(* Logix 5000 project; controller _GigaDiscovery vendor 1 type 14 code 244 rev 35.11; software revision 35.03; part 11 of 23 *)
(* tags used below, declared in another part *)
   Emergencies_CL1 : DINT[14];
(* S_Alarms, continued *)

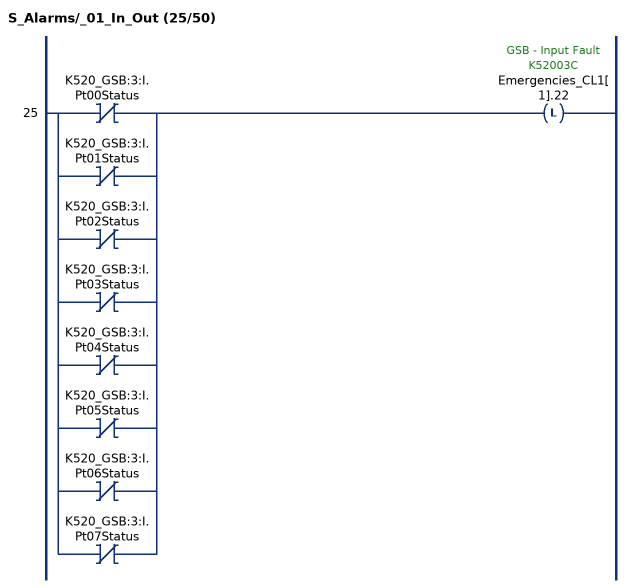
   [picture p185: S_Alarms/_01_In_Out rungs 25-25]
   25: [XIO(K520_GSB:3:I.Pt00Status) ,XIO(K520_GSB:3:I.Pt01Status) ,XIO(K520_GSB:3:I.Pt02Status) ,XIO(K520_GSB:3:I.Pt03Status) ,XIO(K520_GSB:3:I.Pt04Status) ,XIO(K520_GSB:3:I.Pt05Status) ,XIO(K520_GSB:3:I.Pt06Status) ,XIO(K520_GSB:3:I.Pt07Status) ]OTL(Emergencies_CL1[1].22);
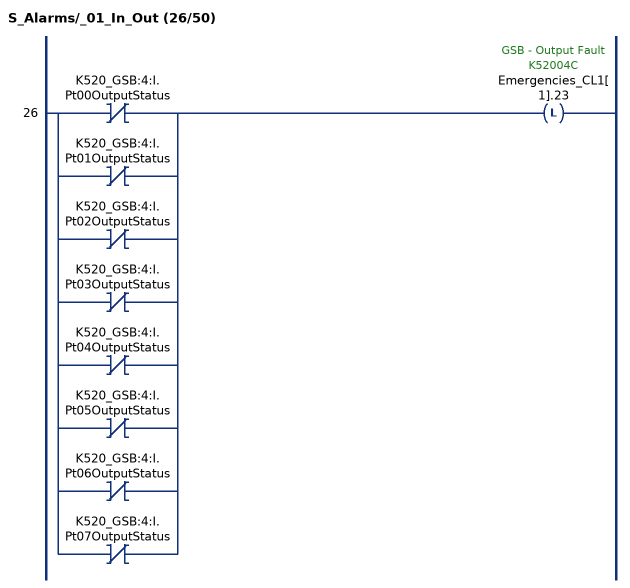
   26: [XIO(K520_GSB:4:I.Pt00OutputStatus) ,XIO(K520_GSB:4:I.Pt01OutputStatus) ,XIO(K520_GSB:4:I.Pt02OutputStatus) ,XIO(K520_GSB:4:I.Pt03OutputStatus) ,XIO(K520_GSB:4:I.Pt04OutputStatus) ,XIO(K520_GSB:4:I.Pt05OutputStatus) ,XIO(K520_GSB:4:I.Pt06OutputStatus) ,XIO(K520_GSB:4:I.Pt07OutputStatus) ]OTL(Emergencies_CL1[1].23);
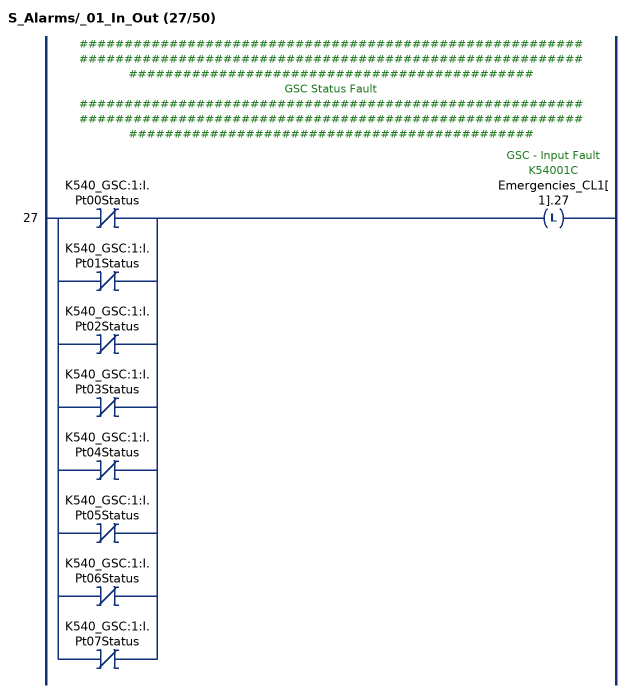
   // #############################################################################################################################################################
   // GSC Status Fault
   // #############################################################################################################################################################
   27: [XIO(K540_GSC:1:I.Pt00Status) ,XIO(K540_GSC:1:I.Pt01Status) ,XIO(K540_GSC:1:I.Pt02Status) ,XIO(K540_GSC:1:I.Pt03Status) ,XIO(K540_GSC:1:I.Pt04Status) ,XIO(K540_GSC:1:I.Pt05Status) ,XIO(K540_GSC:1:I.Pt06Status) ,XIO(K540_GSC:1:I.Pt07Status) ]OTL(Emergencies_CL1[1].27);
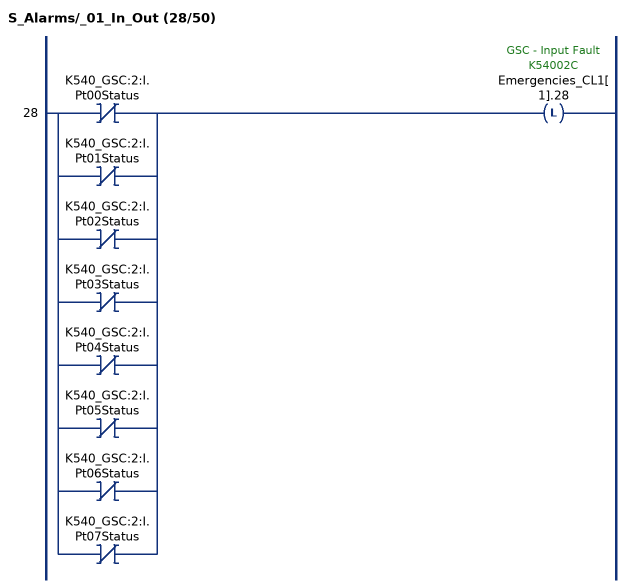
   28: [XIO(K540_GSC:2:I.Pt00Status) ,XIO(K540_GSC:2:I.Pt01Status) ,XIO(K540_GSC:2:I.Pt02Status) ,XIO(K540_GSC:2:I.Pt03Status) ,XIO(K540_GSC:2:I.Pt04Status) ,XIO(K540_GSC:2:I.Pt05Status) ,XIO(K540_GSC:2:I.Pt06Status) ,XIO(K540_GSC:2:I.Pt07Status) ]OTL(Emergencies_CL1[1].28);
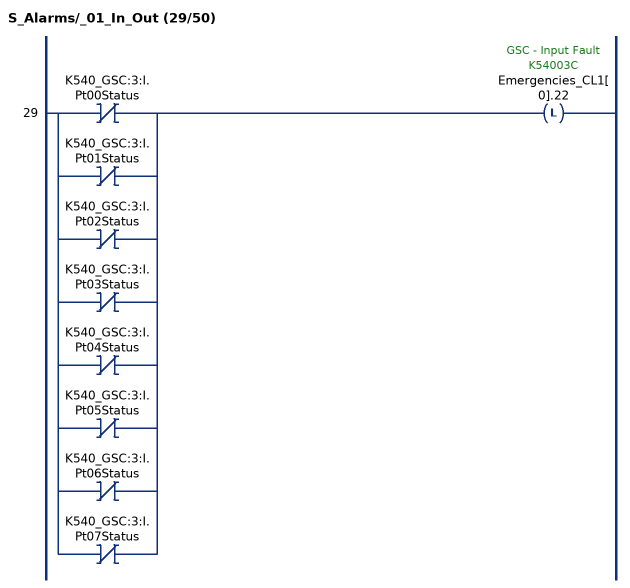
   29: [XIO(K540_GSC:3:I.Pt00Status) ,XIO(K540_GSC:3:I.Pt01Status) ,XIO(K540_GSC:3:I.Pt02Status) ,XIO(K540_GSC:3:I.Pt03Status) ,XIO(K540_GSC:3:I.Pt04Status) ,XIO(K540_GSC:3:I.Pt05Status) ,XIO(K540_GSC:3:I.Pt06Status) ,XIO(K540_GSC:3:I.Pt07Status) ]OTL(Emergencies_CL1[0].22);
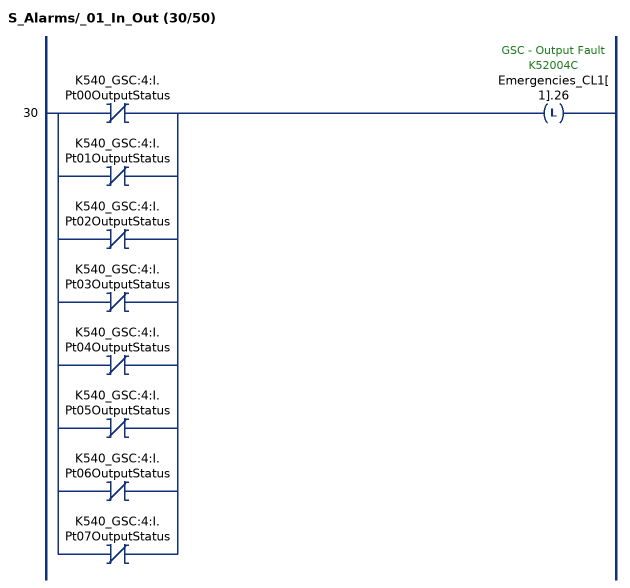
   30: [XIO(K540_GSC:4:I.Pt00OutputStatus) ,XIO(K540_GSC:4:I.Pt01OutputStatus) ,XIO(K540_GSC:4:I.Pt02OutputStatus) ,XIO(K540_GSC:4:I.Pt03OutputStatus) ,XIO(K540_GSC:4:I.Pt04OutputStatus) ,XIO(K540_GSC:4:I.Pt05OutputStatus) ,XIO(K540_GSC:4:I.Pt06OutputStatus) ,XIO(K540_GSC:4:I.Pt07OutputStatus) ]OTL(Emergencies_CL1[1].26);
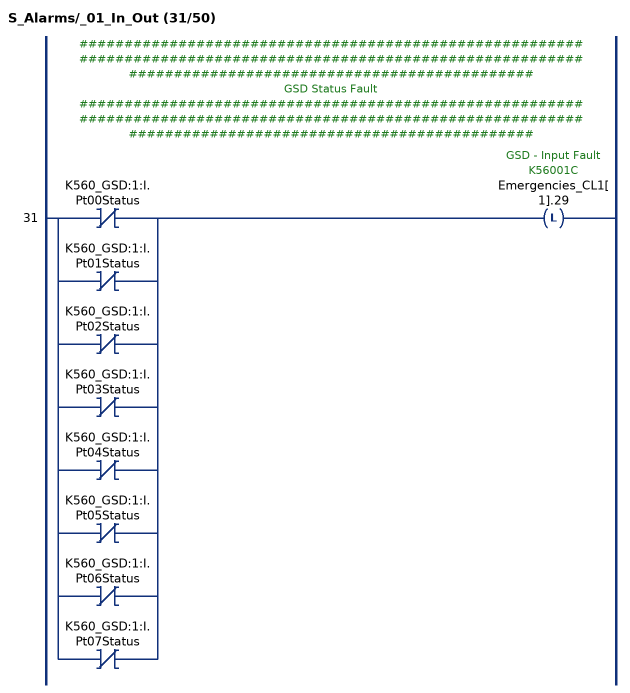
   // #############################################################################################################################################################
   // GSD Status Fault
   // #############################################################################################################################################################
   31: [XIO(K560_GSD:1:I.Pt00Status) ,XIO(K560_GSD:1:I.Pt01Status) ,XIO(K560_GSD:1:I.Pt02Status) ,XIO(K560_GSD:1:I.Pt03Status) ,XIO(K560_GSD:1:I.Pt04Status) ,XIO(K560_GSD:1:I.Pt05Status) ,XIO(K560_GSD:1:I.Pt06Status) ,XIO(K560_GSD:1:I.Pt07Status) ]OTL(Emergencies_CL1[1].29);
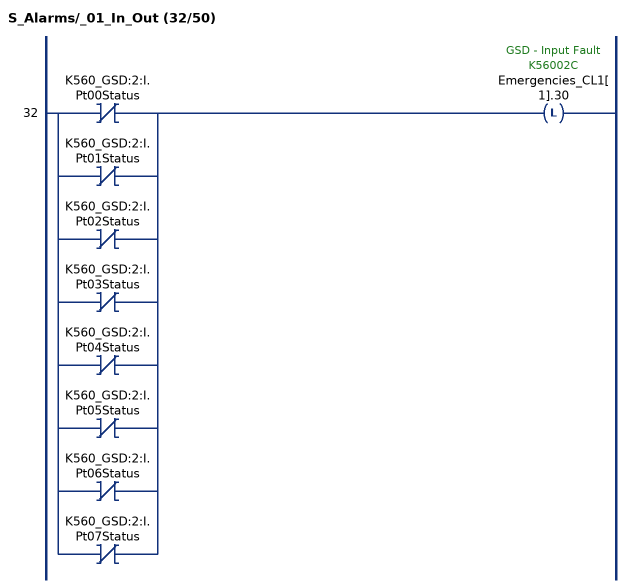
   32: [XIO(K560_GSD:2:I.Pt00Status) ,XIO(K560_GSD:2:I.Pt01Status) ,XIO(K560_GSD:2:I.Pt02Status) ,XIO(K560_GSD:2:I.Pt03Status) ,XIO(K560_GSD:2:I.Pt04Status) ,XIO(K560_GSD:2:I.Pt05Status) ,XIO(K560_GSD:2:I.Pt06Status) ,XIO(K560_GSD:2:I.Pt07Status) ]OTL(Emergencies_CL1[1].30);
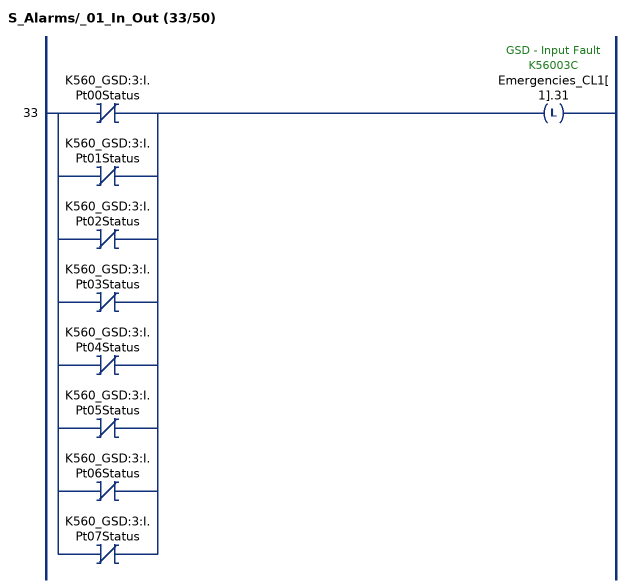
   33: [XIO(K560_GSD:3:I.Pt00Status) ,XIO(K560_GSD:3:I.Pt01Status) ,XIO(K560_GSD:3:I.Pt02Status) ,XIO(K560_GSD:3:I.Pt03Status) ,XIO(K560_GSD:3:I.Pt04Status) ,XIO(K560_GSD:3:I.Pt05Status) ,XIO(K560_GSD:3:I.Pt06Status) ,XIO(K560_GSD:3:I.Pt07Status) ]OTL(Emergencies_CL1[1].31);
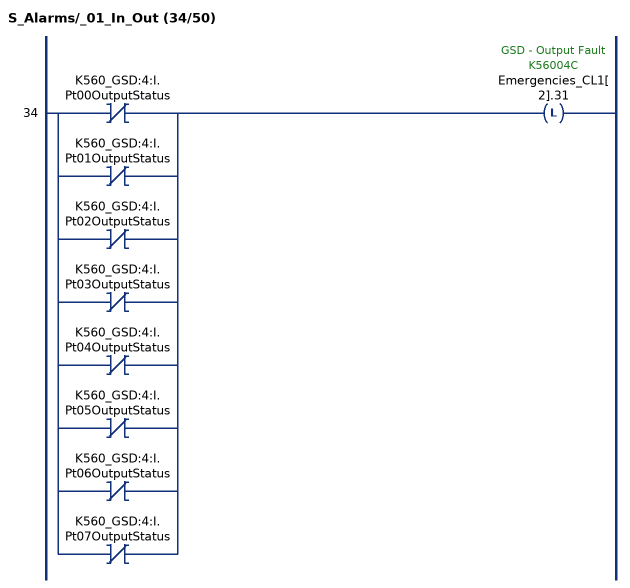
   34: [XIO(K560_GSD:4:I.Pt00OutputStatus) ,XIO(K560_GSD:4:I.Pt01OutputStatus) ,XIO(K560_GSD:4:I.Pt02OutputStatus) ,XIO(K560_GSD:4:I.Pt03OutputStatus) ,XIO(K560_GSD:4:I.Pt04OutputStatus) ,XIO(K560_GSD:4:I.Pt05OutputStatus) ,XIO(K560_GSD:4:I.Pt06OutputStatus) ,XIO(K560_GSD:4:I.Pt07OutputStatus) ]OTL(Emergencies_CL1[2].31);
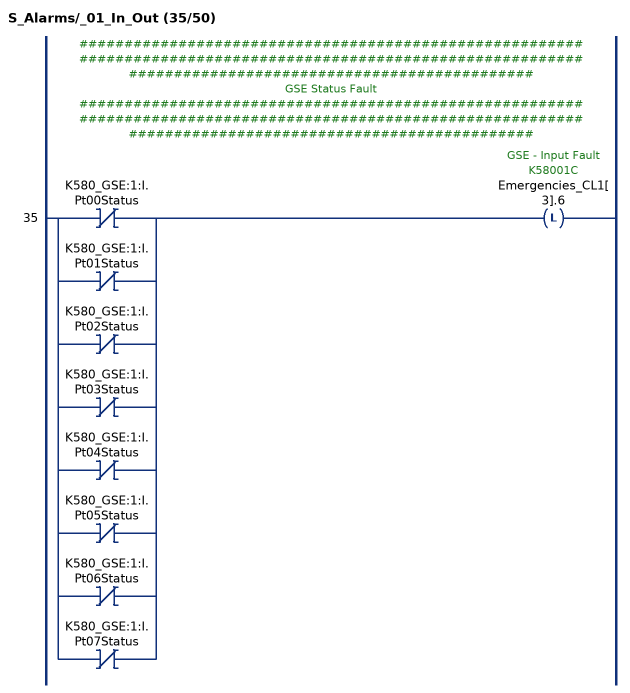
   // #############################################################################################################################################################
   // GSE Status Fault
   // #############################################################################################################################################################
   35: [XIO(K580_GSE:1:I.Pt00Status) ,XIO(K580_GSE:1:I.Pt01Status) ,XIO(K580_GSE:1:I.Pt02Status) ,XIO(K580_GSE:1:I.Pt03Status) ,XIO(K580_GSE:1:I.Pt04Status) ,XIO(K580_GSE:1:I.Pt05Status) ,XIO(K580_GSE:1:I.Pt06Status) ,XIO(K580_GSE:1:I.Pt07Status) ]OTL(Emergencies_CL1[3].6);
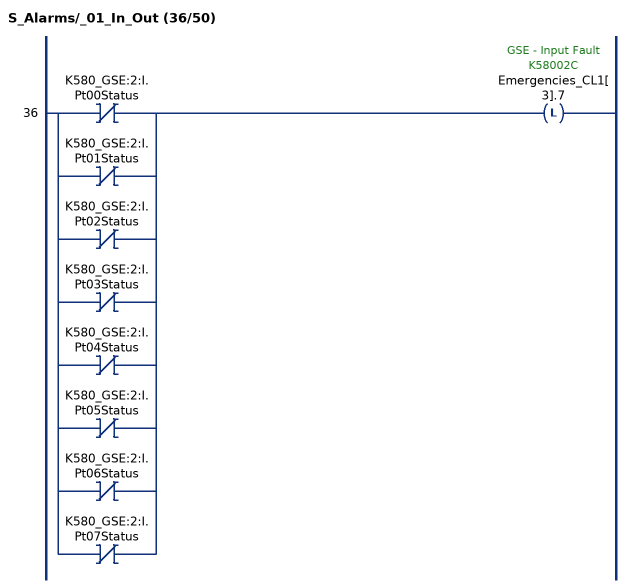
   36: [XIO(K580_GSE:2:I.Pt00Status) ,XIO(K580_GSE:2:I.Pt01Status) ,XIO(K580_GSE:2:I.Pt02Status) ,XIO(K580_GSE:2:I.Pt03Status) ,XIO(K580_GSE:2:I.Pt04Status) ,XIO(K580_GSE:2:I.Pt05Status) ,XIO(K580_GSE:2:I.Pt06Status) ,XIO(K580_GSE:2:I.Pt07Status) ]OTL(Emergencies_CL1[3].7);
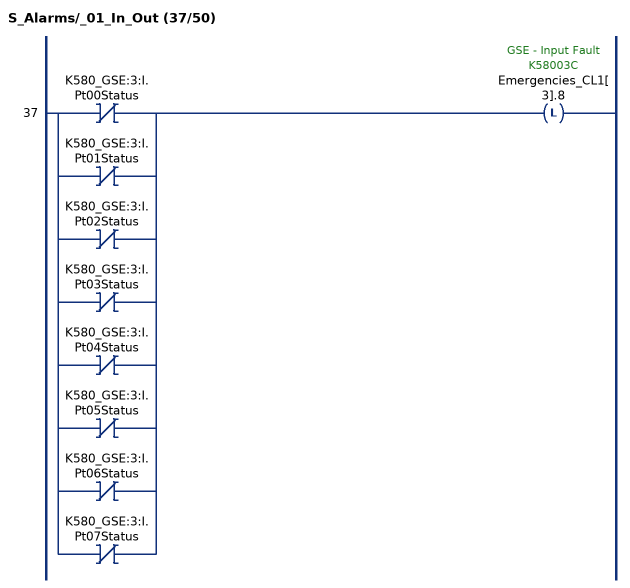
   37: [XIO(K580_GSE:3:I.Pt00Status) ,XIO(K580_GSE:3:I.Pt01Status) ,XIO(K580_GSE:3:I.Pt02Status) ,XIO(K580_GSE:3:I.Pt03Status) ,XIO(K580_GSE:3:I.Pt04Status) ,XIO(K580_GSE:3:I.Pt05Status) ,XIO(K580_GSE:3:I.Pt06Status) ,XIO(K580_GSE:3:I.Pt07Status) ]OTL(Emergencies_CL1[3].8);
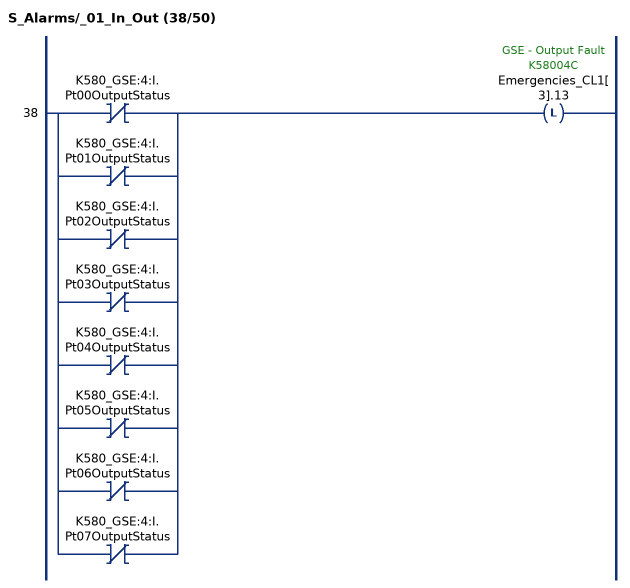
   38: [XIO(K580_GSE:4:I.Pt00OutputStatus) ,XIO(K580_GSE:4:I.Pt01OutputStatus) ,XIO(K580_GSE:4:I.Pt02OutputStatus) ,XIO(K580_GSE:4:I.Pt03OutputStatus) ,XIO(K580_GSE:4:I.Pt04OutputStatus) ,XIO(K580_GSE:4:I.Pt05OutputStatus) ,XIO(K580_GSE:4:I.Pt06OutputStatus) ,XIO(K580_GSE:4:I.Pt07OutputStatus) ]OTL(Emergencies_CL1[3].13);
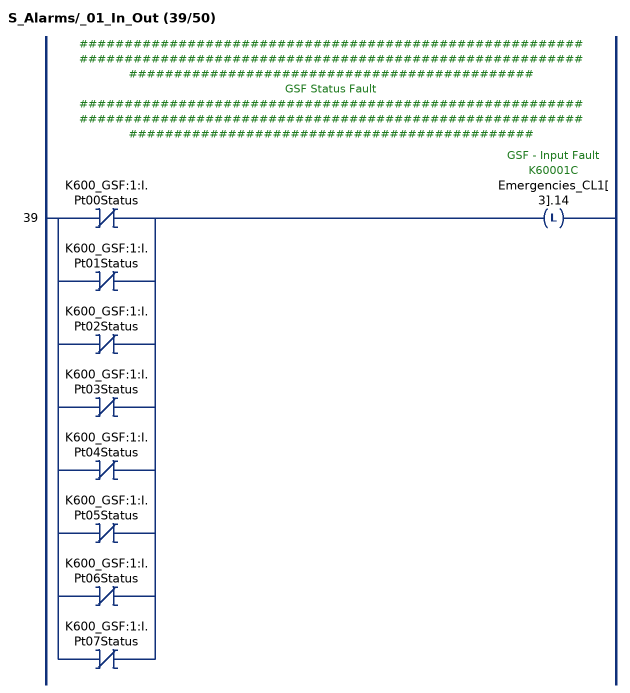
   // #############################################################################################################################################################
   // GSF Status Fault
   // #############################################################################################################################################################
   39: [XIO(K600_GSF:1:I.Pt00Status) ,XIO(K600_GSF:1:I.Pt01Status) ,XIO(K600_GSF:1:I.Pt02Status) ,XIO(K600_GSF:1:I.Pt03Status) ,XIO(K600_GSF:1:I.Pt04Status) ,XIO(K600_GSF:1:I.Pt05Status) ,XIO(K600_GSF:1:I.Pt06Status) ,XIO(K600_GSF:1:I.Pt07Status) ]OTL(Emergencies_CL1[3].14);
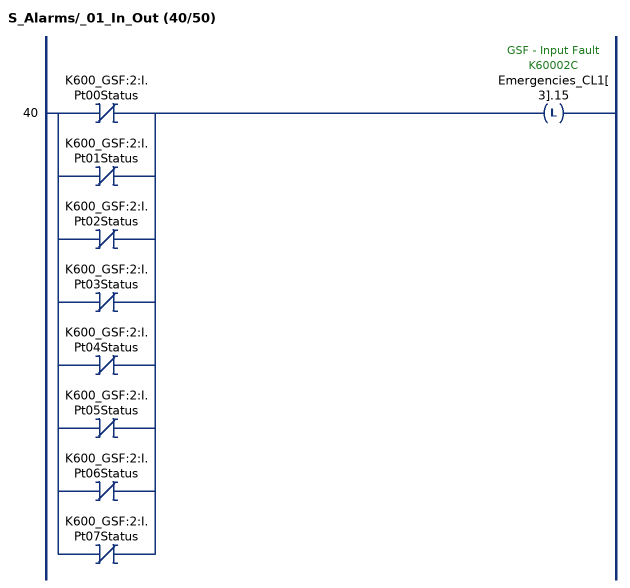
   40: [XIO(K600_GSF:2:I.Pt00Status) ,XIO(K600_GSF:2:I.Pt01Status) ,XIO(K600_GSF:2:I.Pt02Status) ,XIO(K600_GSF:2:I.Pt03Status) ,XIO(K600_GSF:2:I.Pt04Status) ,XIO(K600_GSF:2:I.Pt05Status) ,XIO(K600_GSF:2:I.Pt06Status) ,XIO(K600_GSF:2:I.Pt07Status) ]OTL(Emergencies_CL1[3].15);
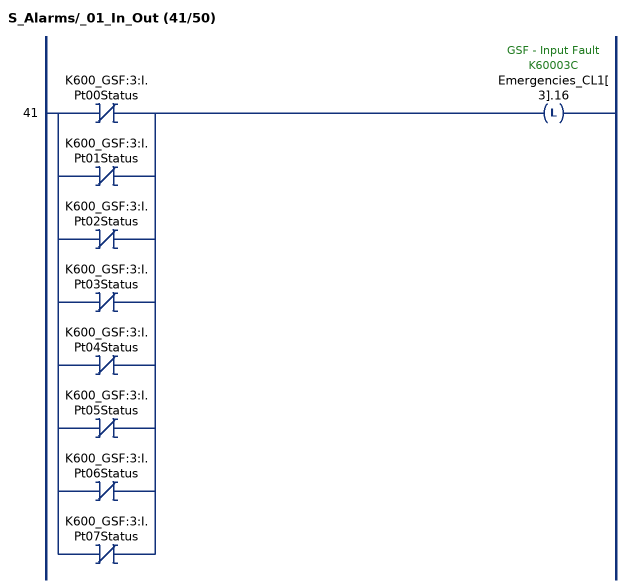
   41: [XIO(K600_GSF:3:I.Pt00Status) ,XIO(K600_GSF:3:I.Pt01Status) ,XIO(K600_GSF:3:I.Pt02Status) ,XIO(K600_GSF:3:I.Pt03Status) ,XIO(K600_GSF:3:I.Pt04Status) ,XIO(K600_GSF:3:I.Pt05Status) ,XIO(K600_GSF:3:I.Pt06Status) ,XIO(K600_GSF:3:I.Pt07Status) ]OTL(Emergencies_CL1[3].16);
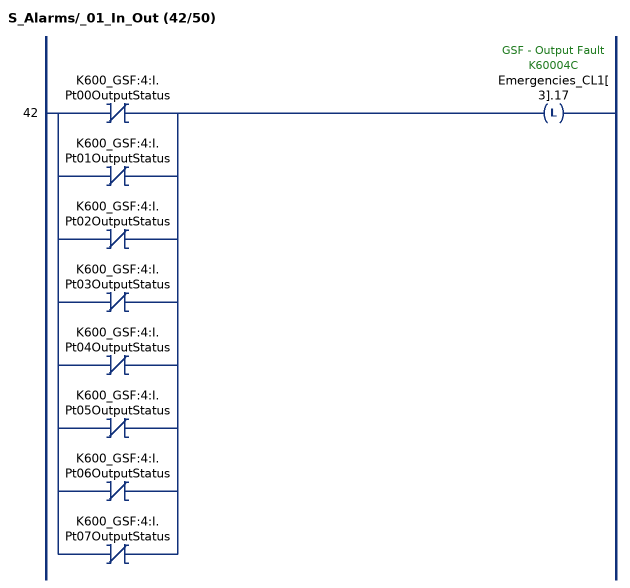
   42: [XIO(K600_GSF:4:I.Pt00OutputStatus) ,XIO(K600_GSF:4:I.Pt01OutputStatus) ,XIO(K600_GSF:4:I.Pt02OutputStatus) ,XIO(K600_GSF:4:I.Pt03OutputStatus) ,XIO(K600_GSF:4:I.Pt04OutputStatus) ,XIO(K600_GSF:4:I.Pt05OutputStatus) ,XIO(K600_GSF:4:I.Pt06OutputStatus) ,XIO(K600_GSF:4:I.Pt07OutputStatus) ]OTL(Emergencies_CL1[3].17);
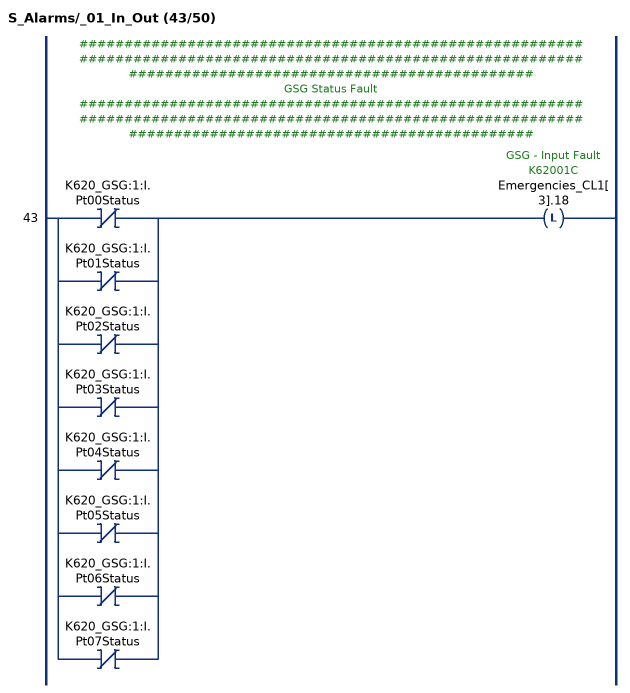
   // #############################################################################################################################################################
   // GSG Status Fault
   // #############################################################################################################################################################
   43: [XIO(K620_GSG:1:I.Pt00Status) ,XIO(K620_GSG:1:I.Pt01Status) ,XIO(K620_GSG:1:I.Pt02Status) ,XIO(K620_GSG:1:I.Pt03Status) ,XIO(K620_GSG:1:I.Pt04Status) ,XIO(K620_GSG:1:I.Pt05Status) ,XIO(K620_GSG:1:I.Pt06Status) ,XIO(K620_GSG:1:I.Pt07Status) ]OTL(Emergencies_CL1[3].18);
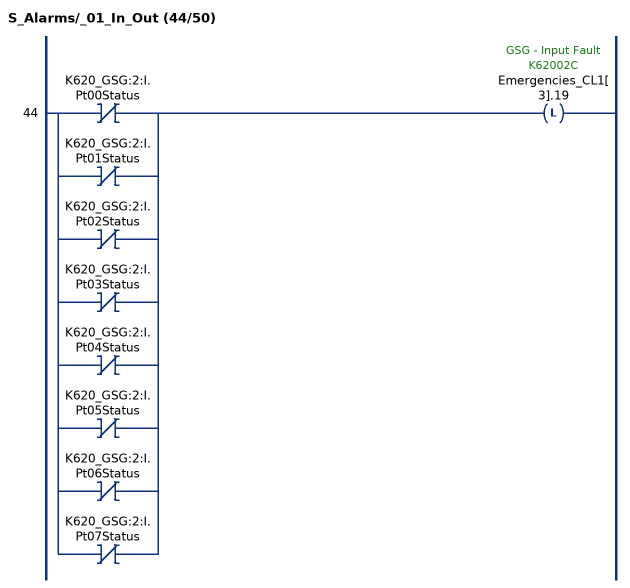
   44: [XIO(K620_GSG:2:I.Pt00Status) ,XIO(K620_GSG:2:I.Pt01Status) ,XIO(K620_GSG:2:I.Pt02Status) ,XIO(K620_GSG:2:I.Pt03Status) ,XIO(K620_GSG:2:I.Pt04Status) ,XIO(K620_GSG:2:I.Pt05Status) ,XIO(K620_GSG:2:I.Pt06Status) ,XIO(K620_GSG:2:I.Pt07Status) ]OTL(Emergencies_CL1[3].19);
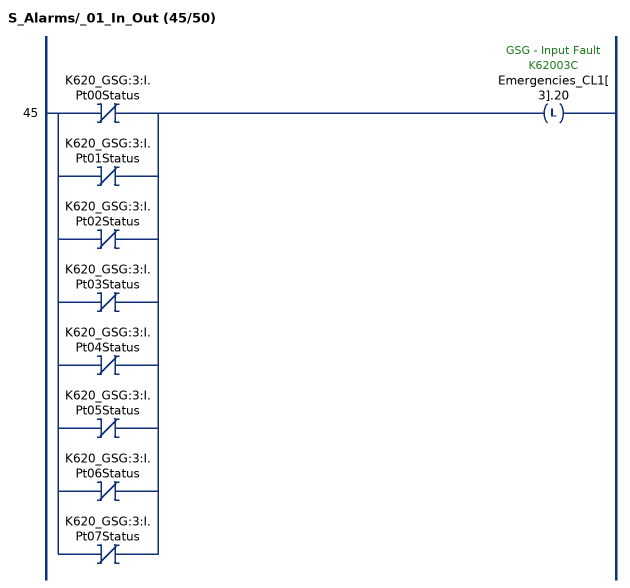
   45: [XIO(K620_GSG:3:I.Pt00Status) ,XIO(K620_GSG:3:I.Pt01Status) ,XIO(K620_GSG:3:I.Pt02Status) ,XIO(K620_GSG:3:I.Pt03Status) ,XIO(K620_GSG:3:I.Pt04Status) ,XIO(K620_GSG:3:I.Pt05Status) ,XIO(K620_GSG:3:I.Pt06Status) ,XIO(K620_GSG:3:I.Pt07Status) ]OTL(Emergencies_CL1[3].20);
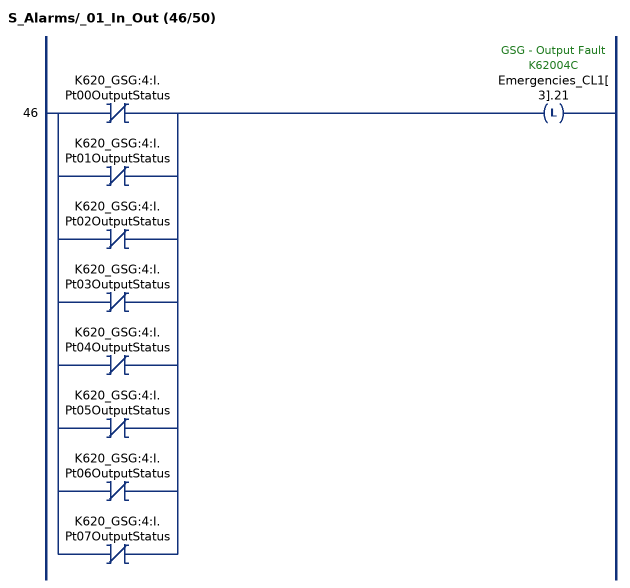
   46: [XIO(K620_GSG:4:I.Pt00OutputStatus) ,XIO(K620_GSG:4:I.Pt01OutputStatus) ,XIO(K620_GSG:4:I.Pt02OutputStatus) ,XIO(K620_GSG:4:I.Pt03OutputStatus) ,XIO(K620_GSG:4:I.Pt04OutputStatus) ,XIO(K620_GSG:4:I.Pt05OutputStatus) ,XIO(K620_GSG:4:I.Pt06OutputStatus) ,XIO(K620_GSG:4:I.Pt07OutputStatus) ]OTL(Emergencies_CL1[3].21);
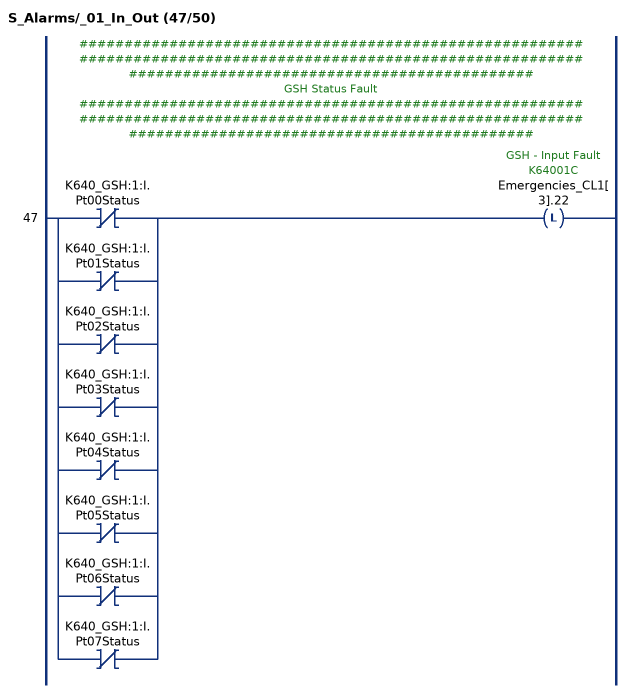
   // #############################################################################################################################################################
   // GSH Status Fault
   // #############################################################################################################################################################
   47: [XIO(K640_GSH:1:I.Pt00Status) ,XIO(K640_GSH:1:I.Pt01Status) ,XIO(K640_GSH:1:I.Pt02Status) ,XIO(K640_GSH:1:I.Pt03Status) ,XIO(K640_GSH:1:I.Pt04Status) ,XIO(K640_GSH:1:I.Pt05Status) ,XIO(K640_GSH:1:I.Pt06Status) ,XIO(K640_GSH:1:I.Pt07Status) ]OTL(Emergencies_CL1[3].22);
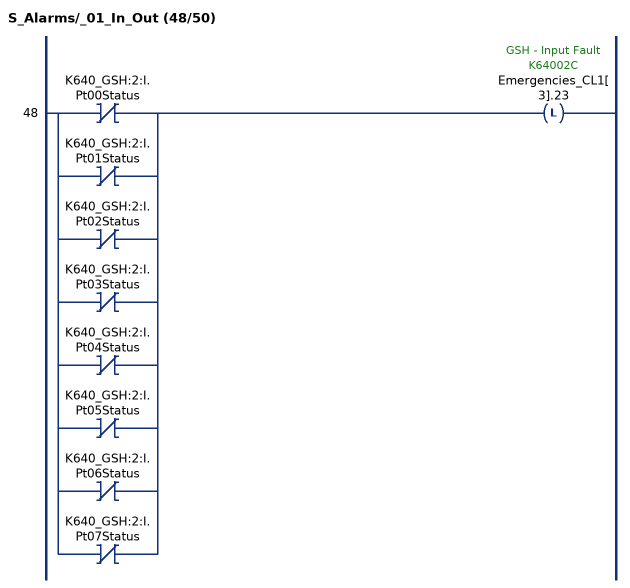
   48: [XIO(K640_GSH:2:I.Pt00Status) ,XIO(K640_GSH:2:I.Pt01Status) ,XIO(K640_GSH:2:I.Pt02Status) ,XIO(K640_GSH:2:I.Pt03Status) ,XIO(K640_GSH:2:I.Pt04Status) ,XIO(K640_GSH:2:I.Pt05Status) ,XIO(K640_GSH:2:I.Pt06Status) ,XIO(K640_GSH:2:I.Pt07Status) ]OTL(Emergencies_CL1[3].23);
